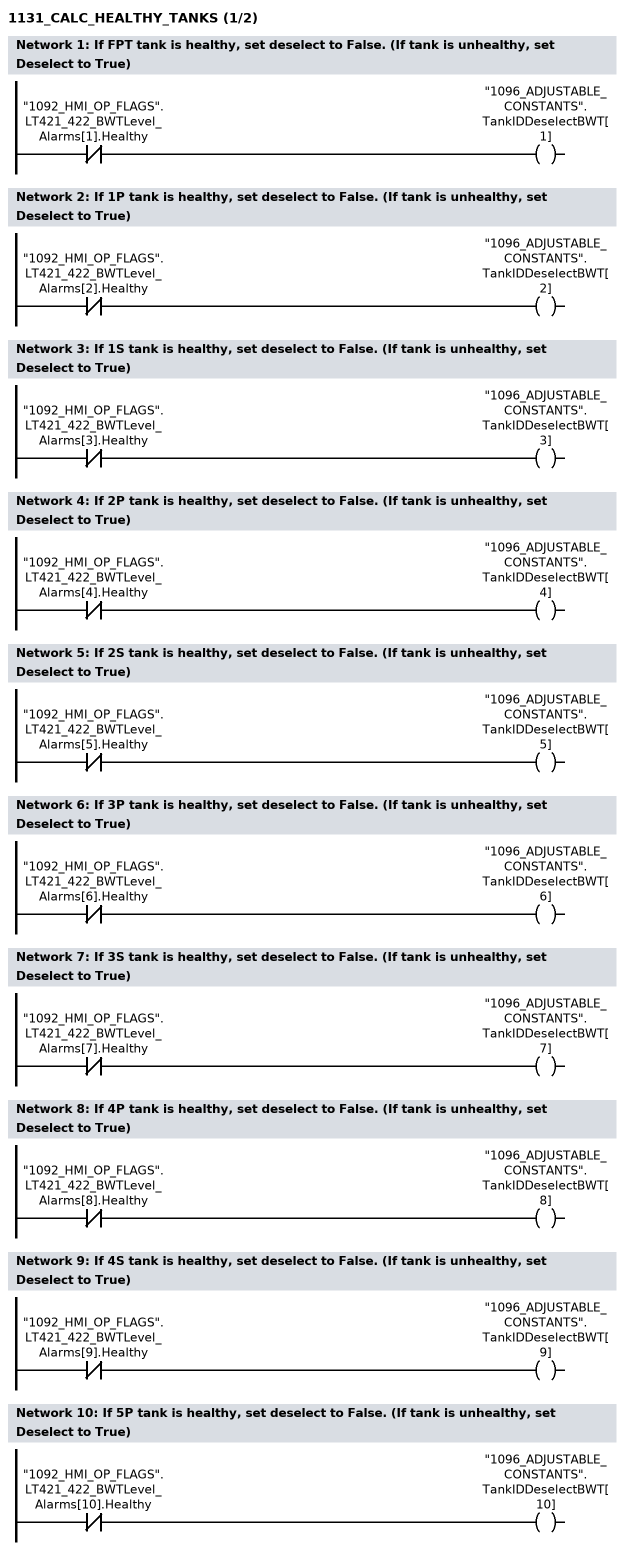
   RUNG wire#powerrail
      I_Contact( "1092_HMI_OP_FLAGS".LT421_422_BWTLevel_Alarms[1].Healthy )
      Coil( "1096_ADJUSTABLE_CONSTANTS".TankIDDeselectBWT[1] )
   END_RUNG
   // the same network as SCL:
   "1096_ADJUSTABLE_CONSTANTS".TankIDDeselectBWT[1] := NOT "1092_HMI_OP_FLAGS".LT421_422_BWTLevel_Alarms[1].Healthy;
END_REGION

REGION Network 2: If 1P tank is healthy, set deselect to False. (If tank is unhealthy, set Deselect to True)
   RUNG wire#powerrail
      I_Contact( "1092_HMI_OP_FLAGS".LT421_422_BWTLevel_Alarms[2].Healthy )
      Coil( "1096_ADJUSTABLE_CONSTANTS".TankIDDeselectBWT[2] )
   END_RUNG
   // the same network as SCL:
   "1096_ADJUSTABLE_CONSTANTS".TankIDDeselectBWT[2] := NOT "1092_HMI_OP_FLAGS".LT421_422_BWTLevel_Alarms[2].Healthy;
END_REGION

REGION Network 3: If 1S tank is healthy, set deselect to False. (If tank is unhealthy, set Deselect to True)
   RUNG wire#powerrail
      I_Contact( "1092_HMI_OP_FLAGS".LT421_422_BWTLevel_Alarms[3].Healthy )
      Coil( "1096_ADJUSTABLE_CONSTANTS".TankIDDeselectBWT[3] )
   END_RUNG
   // the same network as SCL:
   "1096_ADJUSTABLE_CONSTANTS".TankIDDeselectBWT[3] := NOT "1092_HMI_OP_FLAGS".LT421_422_BWTLevel_Alarms[3].Healthy;
END_REGION

REGION Network 4: If 2P tank is healthy, set deselect to False. (If tank is unhealthy, set Deselect to True)
   RUNG wire#powerrail
      I_Contact( "1092_HMI_OP_FLAGS".LT421_422_BWTLevel_Alarms[4].Healthy )
      Coil( "1096_ADJUSTABLE_CONSTANTS".TankIDDeselectBWT[4] )
   END_RUNG
   // the same network as SCL:
   "1096_ADJUSTABLE_CONSTANTS".TankIDDeselectBWT[4] := NOT "1092_HMI_OP_FLAGS".LT421_422_BWTLevel_Alarms[4].Healthy;
END_REGION

REGION Network 5: If 2S tank is healthy, set deselect to False. (If tank is unhealthy, set Deselect to True)
   RUNG wire#powerrail
      I_Contact( "1092_HMI_OP_FLAGS".LT421_422_BWTLevel_Alarms[5].Healthy )
      Coil( "1096_ADJUSTABLE_CONSTANTS".TankIDDeselectBWT[5] )
   END_RUNG
   // the same network as SCL:
   "1096_ADJUSTABLE_CONSTANTS".TankIDDeselectBWT[5] := NOT "1092_HMI_OP_FLAGS".LT421_422_BWTLevel_Alarms[5].Healthy;
END_REGION

REGION Network 6: If 3P tank is healthy, set deselect to False. (If tank is unhealthy, set Deselect to True)
   RUNG wire#powerrail
      I_Contact( "1092_HMI_OP_FLAGS".LT421_422_BWTLevel_Alarms[6].Healthy )
      Coil( "1096_ADJUSTABLE_CONSTANTS".TankIDDeselectBWT[6] )
   END_RUNG
   // the same network as SCL:
   "1096_ADJUSTABLE_CONSTANTS".TankIDDeselectBWT[6] := NOT "1092_HMI_OP_FLAGS".LT421_422_BWTLevel_Alarms[6].Healthy;
END_REGION

REGION Network 7: If 3S tank is healthy, set deselect to False. (If tank is unhealthy, set Deselect to True)
   RUNG wire#powerrail
      I_Contact( "1092_HMI_OP_FLAGS".LT421_422_BWTLevel_Alarms[7].Healthy )
      Coil( "1096_ADJUSTABLE_CONSTANTS".TankIDDeselectBWT[7] )
   END_RUNG
   // the same network as SCL:
   "1096_ADJUSTABLE_CONSTANTS".TankIDDeselectBWT[7] := NOT "1092_HMI_OP_FLAGS".LT421_422_BWTLevel_Alarms[7].Healthy;
END_REGION

REGION Network 8: If 4P tank is healthy, set deselect to False. (If tank is unhealthy, set Deselect to True)
   RUNG wire#powerrail
      I_Contact( "1092_HMI_OP_FLAGS".LT421_422_BWTLevel_Alarms[8].Healthy )
      Coil( "1096_ADJUSTABLE_CONSTANTS".TankIDDeselectBWT[8] )
   END_RUNG
   // the same network as SCL:
   "1096_ADJUSTABLE_CONSTANTS".TankIDDeselectBWT[8] := NOT "1092_HMI_OP_FLAGS".LT421_422_BWTLevel_Alarms[8].Healthy;
END_REGION

REGION Network 9: If 4S tank is healthy, set deselect to False. (If tank is unhealthy, set Deselect to True)
   RUNG wire#powerrail
      I_Contact( "1092_HMI_OP_FLAGS".LT421_422_BWTLevel_Alarms[9].Healthy )
      Coil( "1096_ADJUSTABLE_CONSTANTS".TankIDDeselectBWT[9] )
   END_RUNG
   // the same network as SCL:
   "1096_ADJUSTABLE_CONSTANTS".TankIDDeselectBWT[9] := NOT "1092_HMI_OP_FLAGS".LT421_422_BWTLevel_Alarms[9].Healthy;
END_REGION

REGION Network 10: If 5P tank is healthy, set deselect to False. (If tank is unhealthy, set Deselect to True)
   RUNG wire#powerrail
      I_Contact( "1092_HMI_OP_FLAGS".LT421_422_BWTLevel_Alarms[10].Healthy )
      Coil( "1096_ADJUSTABLE_CONSTANTS".TankIDDeselectBWT[10] )
   END_RUNG
   // the same network as SCL:
   "1096_ADJUSTABLE_CONSTANTS".TankIDDeselectBWT[10] := NOT "1092_HMI_OP_FLAGS".LT421_422_BWTLevel_Alarms[10].Healthy;
END_REGION

REGION Network 11: If 5S tank is healthy, set deselect to False. (If tank is unhealthy, set Deselect to True)
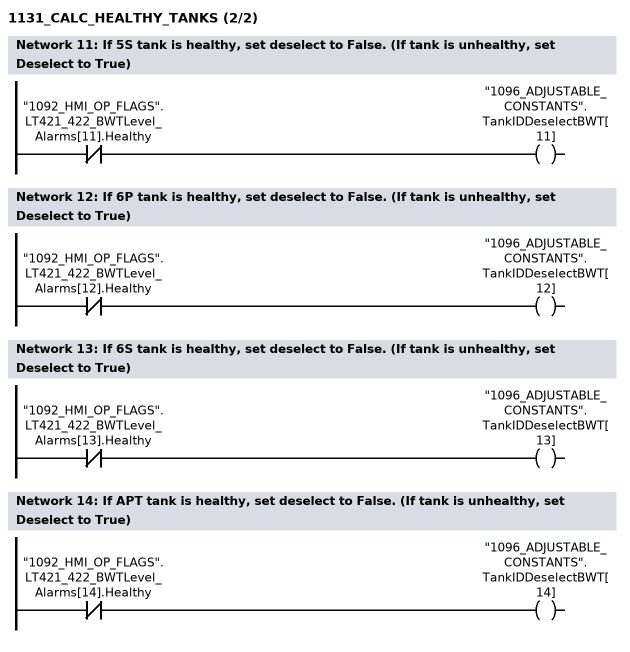
   RUNG wire#powerrail
      I_Contact( "1092_HMI_OP_FLAGS".LT421_422_BWTLevel_Alarms[11].Healthy )
      Coil( "1096_ADJUSTABLE_CONSTANTS".TankIDDeselectBWT[11] )
   END_RUNG
   // the same network as SCL:
   "1096_ADJUSTABLE_CONSTANTS".TankIDDeselectBWT[11] := NOT "1092_HMI_OP_FLAGS".LT421_422_BWTLevel_Alarms[11].Healthy;
END_REGION

REGION Network 12: If 6P tank is healthy, set deselect to False. (If tank is unhealthy, set Deselect to True)
   RUNG wire#powerrail
      I_Contact( "1092_HMI_OP_FLAGS".LT421_422_BWTLevel_Alarms[12].Healthy )
      Coil( "1096_ADJUSTABLE_CONSTANTS".TankIDDeselectBWT[12] )
   END_RUNG
   // the same network as SCL:
   "1096_ADJUSTABLE_CONSTANTS".TankIDDeselectBWT[12] := NOT "1092_HMI_OP_FLAGS".LT421_422_BWTLevel_Alarms[12].Healthy;
END_REGION

REGION Network 13: If 6S tank is healthy, set deselect to False. (If tank is unhealthy, set Deselect to True)
   RUNG wire#powerrail
      I_Contact( "1092_HMI_OP_FLAGS".LT421_422_BWTLevel_Alarms[13].Healthy )
      Coil( "1096_ADJUSTABLE_CONSTANTS".TankIDDeselectBWT[13] )
   END_RUNG
   // the same network as SCL:
   "1096_ADJUSTABLE_CONSTANTS".TankIDDeselectBWT[13] := NOT "1092_HMI_OP_FLAGS".LT421_422_BWTLevel_Alarms[13].Healthy;
END_REGION

REGION Network 14: If APT tank is healthy, set deselect to False. (If tank is unhealthy, set Deselect to True)
   RUNG wire#powerrail
      I_Contact( "1092_HMI_OP_FLAGS".LT421_422_BWTLevel_Alarms[14].Healthy )
      Coil( "1096_ADJUSTABLE_CONSTANTS".TankIDDeselectBWT[14] )
   END_RUNG
   // the same network as SCL:
   "1096_ADJUSTABLE_CONSTANTS".TankIDDeselectBWT[14] := NOT "1092_HMI_OP_FLAGS".LT421_422_BWTLevel_Alarms[14].Healthy;
END_REGION
END_FUNCTION

FUNCTION "1132_CALC_ACTIVE_TANKS" : Void   // FC1132, SCL
{ S7_Optimized_Access := 'TRUE' }
VERSION : 0.1
   VAR_TEMP
      Index : Int;
      NumberActiveTanks : Int;
   END_VAR
   VAR CONSTANT
      NumberOfTanks : Int := 14;
   END_VAR
BEGIN
   (*
       Calculate the number OF active tanks. With this data determine the HMI O/P flags:
       1. NoTanksActive (if no tanks are actively selected or healthy)
       2. The treatment time (the total treatment time of the vessel)
       3. Start IGG Warning Time (time flag to base IGG warnings on)
       4. VoyageLessThanTreatmentTime (error flag is the voyage will not be long enough to treat the tanks).
   *)

   #NumberActiveTanks := 0;

   FOR #Index := 1 TO #NumberOfTanks DO
       // For each tank that is not deselectable, force it to be active.
       IF NOT ("1096_ADJUSTABLE_CONSTANTS".TankIDDeselectBWT[#Index]) THEN
           "1096_ADJUSTABLE_CONSTANTS".TankIDActive[#Index] := TRUE;

       END_IF;
       // Check number of active tanks (either set in HMI, or by force above).
       IF "1096_ADJUSTABLE_CONSTANTS".TankIDActive[#Index] THEN
           #NumberActiveTanks += 1;
       END_IF;
   END_FOR;
   "1191_SYSTEM_VARIABLES".NumberOfActiveTanks := #NumberActiveTanks;

   // Push the no tanks active flag if calculated above.
   IF #NumberActiveTanks = 0 THEN
       "1092_HMI_OP_FLAGS".NoTanksActive := TRUE;
   ELSE
       "1092_HMI_OP_FLAGS".NoTanksActive := FALSE;
   END_IF;
END_FUNCTION

FUNCTION "1133_GTT_DETERMINE_EXCLUSIVITY" : Void   // FC1133, SCL
{ S7_Optimized_Access := 'TRUE' }
VERSION : 0.1
   VAR_INPUT
      TankID_InOperation : Int;
      DemandComplete : Bool;
   END_VAR
   VAR_IN_OUT
      GTT_Exclusivity : "GTT_EXCLUSIVITY";
   END_VAR
BEGIN
   (*
       Verify if the demand has been completed. If the demand is not yet complete,
       then keep this tank 'exclusive', i.e. do not allow another tank ID to begin 
       operating its GTT valve until this demand complete signal becomes True.
   *)

   IF NOT #DemandComplete THEN
       #GTT_Exclusivity.Tank_Exclusivity := TRUE;
       #GTT_Exclusivity.TankID_InOperation := #TankID_InOperation;
   ELSE
       #GTT_Exclusivity.Tank_Exclusivity := FALSE;
       #GTT_Exclusivity.TankID_InOperation := 0;
   END_IF;
END_FUNCTION

FUNCTION "1134_MOVE_TANKS_INGROUP_NEW_STATE" : Void   // FC1134, SCL
{ S7_Optimized_Access := 'TRUE' }
VERSION : 0.1
   VAR_INPUT
      State : "SYSTEM_STATES";
      NewState : Int;
   END_VAR
   VAR_IN_OUT
      TankData : Array[1..#NumberOfTanks] of "TANK_DATA";
   END_VAR
   VAR_TEMP
      Index : Int;
   END_VAR
   VAR CONSTANT
      NumberOfTanks : Int := 14;
   END_VAR
BEGIN
   (*
       For each tank, if it's in the current treatment group, 
       move it into the provided "NewState" state.
   *)
   FOR #Index := 1 TO #NumberOfTanks DO
       IF #TankData[#Index].AllocatedTreatmentGroup = #State.TreatmentGroup AND #TankData[#Index].Active THEN
           #TankData[#Index].TankState := #NewState;
       END_IF;
   END_FOR;
END_FUNCTION

FUNCTION "1135_VALVE_OPEN_CLOSE_TIME_SEL" : Time   // FC1135, SCL
{ S7_Optimized_Access := 'TRUE' }
VERSION : 0.1
   VAR_INPUT
      ValveType : Int;   // Valve Type. {0:NC,1:NO}
      ValveDemand : Bool;
      OpenTime : Time;
      CloseTime : Time;
   END_VAR
   VAR_TEMP
      SelectedTime : Time;
   END_VAR
   VAR CONSTANT
      Valve_NormallyClosed : Int := 0;
      Valve_NormallyOpen : Int := 1;
      Demand_Normal : Int := 0;
      Demand_Enable : Int := 1;
   END_VAR
BEGIN
   // Return the correct time for valve openning or closing based on whether
   // the valve is of type "Normally Open" or "Normally Closed" along with the
   // demand on the valve.
   CASE #ValveType OF
       #Valve_NormallyClosed:
           CASE BOOL_TO_INT(#ValveDemand) OF
               #Demand_Normal:
                   #SelectedTime := #CloseTime;
               #Demand_Enable:
                   #SelectedTime := #OpenTime;
           END_CASE;
       #Valve_NormallyOpen:
           CASE BOOL_TO_INT(#ValveDemand) OF
               #Demand_Normal:
                   #SelectedTime := #OpenTime;
               #Demand_Enable:
                   #SelectedTime := #CloseTime;
           END_CASE;
   END_CASE;

   #"1135_VALVE_OPEN_CLOSE_TIME_SEL" := #SelectedTime;
END_FUNCTION

FUNCTION "1136_CALC_NEXT_TREATMENT_GROUP" : Int   // FC1136, SCL
{ S7_Optimized_Access := 'TRUE' }
VERSION : 0.1
   VAR_INPUT
      State : "SYSTEM_STATES";
      NumberOfTreatmentGroups : Int;
      TankData : Array[1..#NumberOfTanks] of "TANK_DATA";
   END_VAR
   VAR_TEMP
      NextTreatmentGroupCalc : Int;
      NextTreatmentGroupFound : Bool;
      TreatmentGroupContainsActiveTank : Bool;
      Index : Int;
   END_VAR
   VAR CONSTANT
      NumberOfTanks : Int := 14;
   END_VAR
BEGIN
   // Return the next treatment group ID which contains active tanks.
   // Return a -1 if there are no further active tanks, or this is the greatest tank ID.
   #NextTreatmentGroupFound := False;
   #NextTreatmentGroupCalc := #State.TreatmentGroup + 1;

   IF #NextTreatmentGroupCalc <= #NumberOfTreatmentGroups THEN
       WHILE NOT #NextTreatmentGroupFound DO
           // Another treatment group to go, check if there are active tanks in the next group.
           #TreatmentGroupContainsActiveTank := False;
           FOR #Index := 1 TO #NumberOfTanks DO
               IF #TankData[#Index].AllocatedTreatmentGroup = #NextTreatmentGroupCalc AND "1096_ADJUSTABLE_CONSTANTS".TankIDActive[#Index] = True THEN
                   #TreatmentGroupContainsActiveTank := True;
               END_IF;
           END_FOR;
           IF #TreatmentGroupContainsActiveTank = True THEN
               // A treatment group has been found.
               #NextTreatmentGroupFound := True;
           ELSE
               // A treatment group was not found on this cycle, check if there are more treatment groups to go.
               IF #NextTreatmentGroupCalc + 1 <= #NumberOfTreatmentGroups THEN
                   #NextTreatmentGroupCalc += 1;
               ELSE
                   // No treatment groups remain, return -1.
                   #NextTreatmentGroupCalc := -1;
                   #NextTreatmentGroupFound := True;
               END_IF;
           END_IF;
       END_WHILE;
   ELSE
       // This is the last treatment group, return a -1 to show that there are no further groups.
       #NextTreatmentGroupCalc := -1;
   END_IF;

   #"1136_CALC_NEXT_TREATMENT_GROUP" := #NextTreatmentGroupCalc;
END_FUNCTION

// folder: 1000 - 1999 BWT System Control/1130 - 1159 Support Functions/1150 - 1159 Next Stage Checks

FUNCTION "1150_NEXT_STAGE_CHECK_GTT" : "ALARM_DEMAND_RTN"   // FC1150, SCL
{ S7_Optimized_Access := 'TRUE' }
VERSION : 0.1
   VAR_INPUT
      AlarmState : Int;   // State system should move to in the event of an alarm being raised (Normally State_Shutdown)
      GTT_OUT : "VALVE_GTT_OUT";
      TankData : Array[1..#NumberOfTanks] of "TANK_DATA";
   END_VAR
   VAR_IN_OUT
      State : "SYSTEM_STATES";
   END_VAR
   VAR_TEMP
      Index : Int;
      NextStageCheck : "ALARM_DEMAND_RTN";
   END_VAR
   VAR CONSTANT
      NumberOfTanks : Int := 14;
   END_VAR
BEGIN
   (*
       Function to check whether the treatment group is ready to move to the next stage
       This specifically checks the GTT completion and will return the demand complete
       only once all active tanks have completed GTT actuation actions.
   *)

   #NextStageCheck.Demand_Complete := True;
   #NextStageCheck.Alarm_Active := False;

   FOR #Index := 1 TO #NumberOfTanks DO
       IF #TankData[#Index].AllocatedTreatmentGroup = #State.TreatmentGroup AND #TankData[#Index].Active THEN
           IF NOT (#GTT_OUT.GTT_DemandsCompleted[#Index]) THEN
               #NextStageCheck.Demand_Complete := False;
           END_IF;
           IF #GTT_OUT.GTT_Alarms[#Index] THEN
               #NextStageCheck.Alarm_Active := True;
           END_IF;
       END_IF;
   END_FOR;

   IF #NextStageCheck.Alarm_Active THEN
       #State.System := #AlarmState;
   END_IF;

   #"1150_NEXT_STAGE_CHECK_GTT" := #NextStageCheck;
END_FUNCTION

FUNCTION "1151_NEXT_STAGE_CHECK_PVV" : "ALARM_DEMAND_RTN"   // FC1151, SCL
{ S7_Optimized_Access := 'TRUE' }
VERSION : 0.1
   VAR_INPUT
      AlarmState : Int;   // State system should move to in the event of an alarm being raised (Normally State_Shutdown)
      PVVX_OUT : "VALVE_PVVX_OUT";
      TankData : Array[1..#NumberOfTanks] of "TANK_DATA";
   END_VAR
   VAR_IN_OUT
      State : "SYSTEM_STATES";
   END_VAR
   VAR_TEMP
      Index : Int;
      NextStageCheck : "ALARM_DEMAND_RTN";
   END_VAR
   VAR CONSTANT
      NumberOfTanks : Int := 14;
   END_VAR
BEGIN
   (*
       Function to check whether the treatment group is ready to move to the next stage
       This specifically checks the Vent A/B completion and will return the demand complete
       only once all active tanks have completed Vent A/B actuation actions.
   *)

   #NextStageCheck.Demand_Complete := True;
   #NextStageCheck.Alarm_Active := False;

   FOR #Index := 1 TO #NumberOfTanks DO
       IF #TankData[#Index].AllocatedTreatmentGroup = #State.TreatmentGroup AND #TankData[#Index].Active THEN
           IF NOT (#PVVX_OUT.PVVA_DemandsCompleted[#Index] OR #PVVX_OUT.PVVB_DemandsCompleted[#Index]) THEN
               #NextStageCheck.Demand_Complete := False;
           END_IF;
           IF (#PVVX_OUT.PVVA_Alarms[#Index] OR #PVVX_OUT.PVVB_Alarms[#Index]) THEN
               #NextStageCheck.Alarm_Active := True;
           END_IF;
       END_IF;
   END_FOR;

   IF #NextStageCheck.Alarm_Active THEN
       #State.System := #AlarmState;
   END_IF;

   #"1151_NEXT_STAGE_CHECK_PVV" := #NextStageCheck;
END_FUNCTION

FUNCTION "1152_NEXT_STAGE_CHECK_TIMER" : "ALARM_DEMAND_RTN"   // FC1152, SCL
{ S7_Optimized_Access := 'TRUE' }
VERSION : 0.1
   VAR_INPUT
      AlarmState : Int;   // State system should move to in the event of an alarm being raised (Normally State_Shutdown)
      TankData : Array[1..#NumberOfTanks] of "TANK_DATA";
   END_VAR
   VAR_IN_OUT
      State : "SYSTEM_STATES";
   END_VAR
   VAR_TEMP
      Index : Int;
      NextStageCheck : "ALARM_DEMAND_RTN";
   END_VAR
   VAR CONSTANT
      NumberOfTanks : Int := 14;
   END_VAR
BEGIN
   (*
       Function to check whether the treatment group is ready to move to the next stage
       This specifically checks the the timer of a tank (xx-Dwell) completion and will return
       the demand complete only once all active tanks have completed their timeouts, depending
       on the overall system state, this is a multi-function block call
   *)

   #NextStageCheck.Demand_Complete := True;
   #NextStageCheck.Alarm_Active := False;

   FOR #Index := 1 TO #NumberOfTanks DO
       IF #TankData[#Index].AllocatedTreatmentGroup = #State.TreatmentGroup AND #TankData[#Index].Active THEN
           IF NOT (#TankData[#Index].Timer_Complete) THEN
               #NextStageCheck.Demand_Complete := False;
           END_IF;
       END_IF;
   END_FOR;

   IF #NextStageCheck.Alarm_Active THEN
       #State.System := #AlarmState;
   END_IF;

   #"1152_NEXT_STAGE_CHECK_TIMER" := #NextStageCheck;
END_FUNCTION

FUNCTION "1153_NEXT_STAGE_CHECK_XEOX" : "ALARM_DEMAND_RTN"   // FC1153, SCL
{ S7_Optimized_Access := 'TRUE' }
VERSION : 0.1
   VAR_INPUT
      AlarmState : Int;   // State system should move to in the event of an alarm being raised (Normally State_Shutdown)
      TankData : Array[1..#NumberOfTanks] of "TANK_DATA";
   END_VAR
   VAR_IN_OUT
      State : "SYSTEM_STATES";
   END_VAR
   VAR_TEMP
      Index : Int;
      NextStageCheck : "ALARM_DEMAND_RTN";
   END_VAR
   VAR CONSTANT
      NumberOfTanks : Int := 14;
   END_VAR
BEGIN
   (*
       Function to check whether the treatment group is ready to move to the next stage
       This specifically checks the the ReOx/DeOx of a tank completion and will return
       the demand complete only once all active tanks have completed ReOx or DeOx, depending
       on the overall system state, this is a multi-function block call
   *)

   #NextStageCheck.Demand_Complete := True;
   #NextStageCheck.Alarm_Active := False;

   FOR #Index := 1 TO #NumberOfTanks DO
       IF #TankData[#Index].AllocatedTreatmentGroup = #State.TreatmentGroup AND #TankData[#Index].Active THEN
           IF NOT (#TankData[#Index].XeOx_Complete) THEN
               #NextStageCheck.Demand_Complete := False;
           END_IF;
       END_IF;
   END_FOR;

   IF #NextStageCheck.Alarm_Active THEN
       #State.System := #AlarmState;
   END_IF;

   #"1153_NEXT_STAGE_CHECK_XEOX" := #NextStageCheck;
END_FUNCTION

// folder: 1000 - 1999 BWT System Control/1600 - 1999 Standard FB's

FUNCTION_BLOCK "1604_DEMAND_AND_CHECK"   // FB1604, LAD
TITLE = Valve Check
{ S7_Optimized_Access := 'TRUE' }
AUTHOR : JRS
VERSION : 0.1
// Demand and check an NO or NC valve.
   VAR_INPUT
      DemandIn : Bool;   // Demand
      NO_Type : Bool;   // Valve type = open without demand
      NC_Type : Bool;   // Valve type = closed without demand
      ValveMoveTime : LTime := LT#1s;   // Maximum movement time
      ValveOpenStatus : Bool;   // Valve open confirmed
      ValveClsdStatus : Bool;   // Valve closed confirmed
   END_VAR
   VAR_OUTPUT
      DemandOut : Bool;   // Demand feedthrough from DemandIn
      DemandComplete : Bool;   // Valve has completed movement
      Alarm : Bool;   // Valve is faulty
   END_VAR
   VAR RETAIN
      Reset : Bool := True;
      Healthy : Bool;   // Valve is healthy
      Config_Error : Bool;   // Configuration error
      Sensor_Fault : Bool;   // Sensor conflicts
      TRAVEL_TIME : TONR_LTIME;
   END_VAR
BEGIN

REGION Network 1: Configuration Error
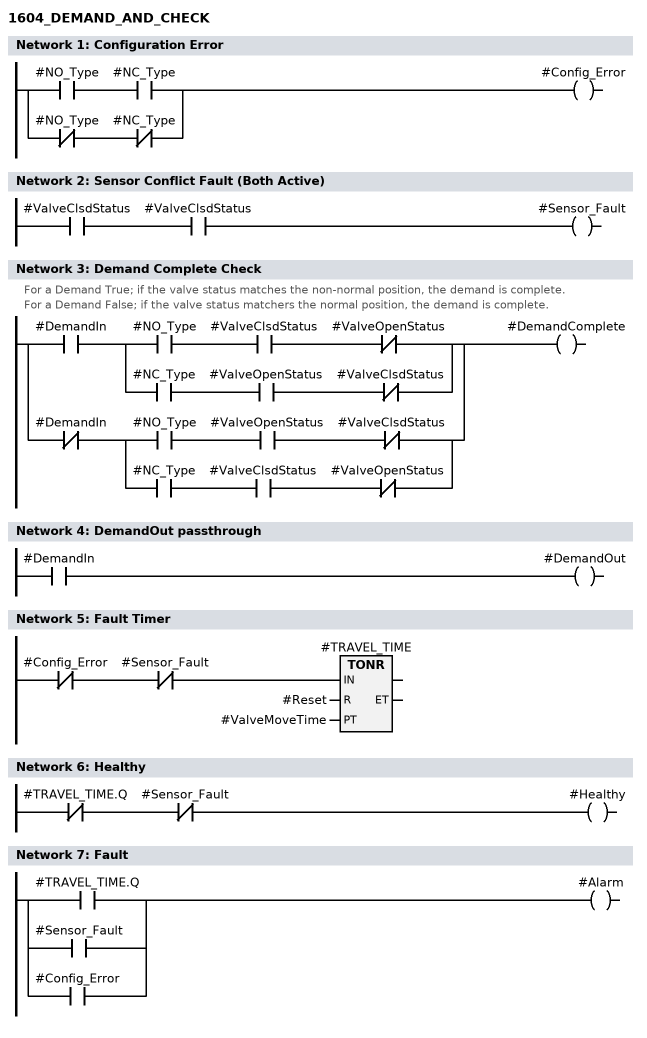
   RUNG wire#powerrail
      Contact( #NO_Type )
      Contact( #NC_Type )
      wire#w1
      Coil( #Config_Error )
   END_RUNG
   RUNG wire#powerrail
      I_Contact( #NO_Type )
      I_Contact( #NC_Type )
   END_RUNG wire#w1
   // the same network as SCL:
   #Config_Error := (#NO_Type AND #NC_Type) OR (NOT #NO_Type AND NOT #NC_Type);
END_REGION

REGION Network 2: Sensor Conflict Fault (Both Active)
   RUNG wire#powerrail
      Contact( #ValveClsdStatus )
      Contact( #ValveClsdStatus )
      Coil( #Sensor_Fault )
   END_RUNG
   // the same network as SCL:
   #Sensor_Fault := #ValveClsdStatus AND #ValveClsdStatus;
END_REGION

REGION Network 3: Demand Complete Check
   // For a Demand True; if the valve status matches the non-normal position, the demand is complete.
   // For a Demand False; if the valve status matchers the normal position, the demand is complete.
   RUNG wire#powerrail
      Contact( #DemandIn )
      wire#w1
      Contact( #NO_Type )
      Contact( #ValveClsdStatus )
      I_Contact( #ValveOpenStatus )
      wire#w2
      Coil( #DemandComplete )
   END_RUNG
   RUNG wire#w1
      Contact( #NC_Type )
      Contact( #ValveOpenStatus )
      I_Contact( #ValveClsdStatus )
   END_RUNG wire#w2
   RUNG wire#powerrail
      I_Contact( #DemandIn )
      wire#w3
      Contact( #NO_Type )
      Contact( #ValveOpenStatus )
      I_Contact( #ValveClsdStatus )
   END_RUNG wire#w2
   RUNG wire#w3
      Contact( #NC_Type )
      Contact( #ValveClsdStatus )
      I_Contact( #ValveOpenStatus )
   END_RUNG wire#w2
   // the same network as SCL:
   #DemandComplete := (#DemandIn AND ((#NO_Type AND #ValveClsdStatus AND NOT #ValveOpenStatus) OR (#NC_Type AND #ValveOpenStatus AND NOT #ValveClsdStatus))) OR (NOT #DemandIn AND ((#NO_Type AND #ValveOpenStatus AND NOT #ValveClsdStatus) OR (#NC_Type AND #ValveClsdStatus AND NOT #ValveOpenStatus)));
END_REGION

REGION Network 4: DemandOut passthrough
   RUNG wire#powerrail
      Contact( #DemandIn )
      Coil( #DemandOut )
   END_RUNG
   // the same network as SCL:
   #DemandOut := #DemandIn;
END_REGION

REGION Network 5: Fault Timer
   #TRAVEL_TIME(IN := NOT #Config_Error AND NOT #Sensor_Fault, R := #Reset, PT := #ValveMoveTime);   // TONR
END_REGION

REGION Network 6: Healthy
   RUNG wire#powerrail
      I_Contact( #TRAVEL_TIME.Q )
      I_Contact( #Sensor_Fault )
      Coil( #Healthy )
   END_RUNG
   // the same network as SCL:
   #Healthy := NOT #TRAVEL_TIME.Q AND NOT #Sensor_Fault;
END_REGION

REGION Network 7: Fault
   RUNG wire#powerrail
      Contact( #TRAVEL_TIME.Q )
      wire#w1
      Coil( #Alarm )
   END_RUNG
   RUNG wire#powerrail
      Contact( #Sensor_Fault )
   END_RUNG wire#w1
   RUNG wire#powerrail
      Contact( #Config_Error )
   END_RUNG wire#w1
   // the same network as SCL:
   #Alarm := #TRAVEL_TIME.Q OR #Sensor_Fault OR #Config_Error;
END_REGION
END_FUNCTION_BLOCK

FUNCTION "1601_ANALOGUE_HEALTH_ALLTRIPS" : Void   // FC1601, LAD
{ S7_Optimized_Access := 'TRUE' }
VERSION : 0.1
   VAR_INPUT
      InputSignal : Real;   // Analogue sensor value
      InputMinimum : Real;   // Minimum sensor value
      InputMaximum : Real;   // Maximum sensor value
      InputSetpointLowLow : Real;   // Low low setpoint value for sensor
      InputSetpointLow : Real;   // Low setpoint value for sensor
      InputSetpointHigh : Real;   // High setpoint value for sensor
      InputSetpointHighHigh : Real;   // High high setpoint value for sensor
   END_VAR
   VAR_OUTPUT
      SensorHealthOut : Bool;   // Boolean health status
      LowLowAlarmOut : Bool;   // Boolean for low low alarm
      LowWarningOut : Bool;   // Boolean for low warning
      HighWarningOut : Bool;   // Boolean for high warning
      HighHighAlarmOut : Bool;   // Boolean for high high alarm
   END_VAR
BEGIN

REGION Network 1: Boolean health status
   // Determine SensorHealthOut (health status) dependent on input signal from sensor compared to setpoints. [GEN-05]
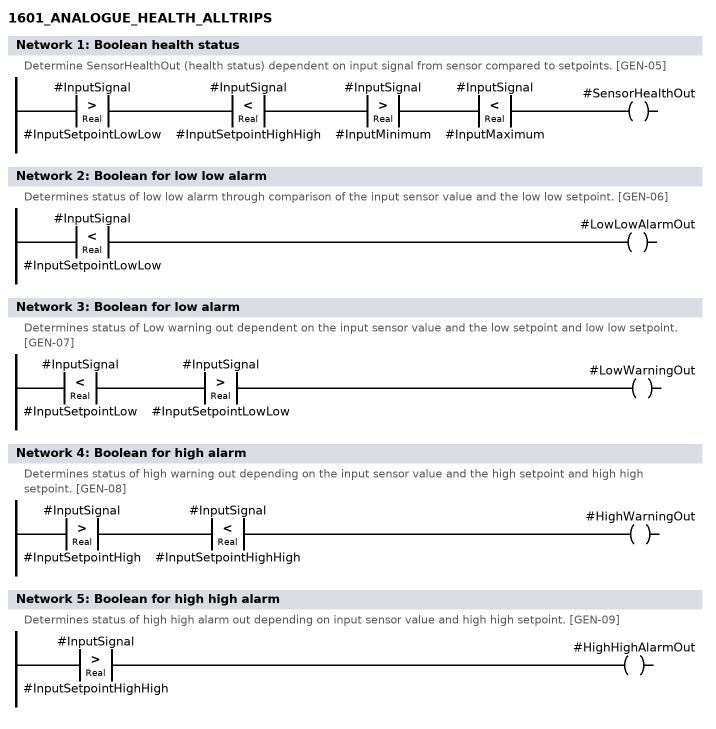
   RUNG wire#powerrail
      { S7_Templates := "SrcType := Real" } GT_Contact(in1 := #InputSignal, in2 := #InputSetpointLowLow)
      { S7_Templates := "SrcType := Real" } LT_Contact(in1 := #InputSignal, in2 := #InputSetpointHighHigh)
      { S7_Templates := "SrcType := Real" } GT_Contact(in1 := #InputSignal, in2 := #InputMinimum)
      { S7_Templates := "SrcType := Real" } LT_Contact(in1 := #InputSignal, in2 := #InputMaximum)
      Coil( #SensorHealthOut )
   END_RUNG
   // the same network as SCL:
   #SensorHealthOut := (#InputSignal > #InputSetpointLowLow) AND (#InputSignal < #InputSetpointHighHigh) AND (#InputSignal > #InputMinimum) AND (#InputSignal < #InputMaximum);
END_REGION

REGION Network 2: Boolean for low low alarm
   // Determines status of low low alarm through comparison of the input sensor value and the low low setpoint. [GEN-06]
   RUNG wire#powerrail
      { S7_Templates := "SrcType := Real" } LT_Contact(in1 := #InputSignal, in2 := #InputSetpointLowLow)
      Coil( #LowLowAlarmOut )
   END_RUNG
   // the same network as SCL:
   #LowLowAlarmOut := #InputSignal < #InputSetpointLowLow;
END_REGION

REGION Network 3: Boolean for low alarm
   // Determines status of Low warning out dependent on the input sensor value and the low setpoint and low low setpoint. [GEN-07]
   RUNG wire#powerrail
      { S7_Templates := "SrcType := Real" } LT_Contact(in1 := #InputSignal, in2 := #InputSetpointLow)
      { S7_Templates := "SrcType := Real" } GT_Contact(in1 := #InputSignal, in2 := #InputSetpointLowLow)
      Coil( #LowWarningOut )
   END_RUNG
   // the same network as SCL:
   #LowWarningOut := (#InputSignal < #InputSetpointLow) AND (#InputSignal > #InputSetpointLowLow);
END_REGION

REGION Network 4: Boolean for high alarm
   // Determines status of high warning out depending on the input sensor value and the high setpoint and high high setpoint. [GEN-08]
   RUNG wire#powerrail
      { S7_Templates := "SrcType := Real" } GT_Contact(in1 := #InputSignal, in2 := #InputSetpointHigh)
      { S7_Templates := "SrcType := Real" } LT_Contact(in1 := #InputSignal, in2 := #InputSetpointHighHigh)
      Coil( #HighWarningOut )
   END_RUNG
   // the same network as SCL:
   #HighWarningOut := (#InputSignal > #InputSetpointHigh) AND (#InputSignal < #InputSetpointHighHigh);
END_REGION

REGION Network 5: Boolean for high high alarm
   // Determines status of high high alarm out depending on input sensor value and high high setpoint. [GEN-09]
   RUNG wire#powerrail
      { S7_Templates := "SrcType := Real" } GT_Contact(in1 := #InputSignal, in2 := #InputSetpointHighHigh)
      Coil( #HighHighAlarmOut )
   END_RUNG
   // the same network as SCL:
   #HighHighAlarmOut := #InputSignal > #InputSetpointHighHigh;
END_REGION
END_FUNCTION

FUNCTION "1602_DIGITAL_HEALTH" : Void   // FC1602, LAD
{ S7_Optimized_Access := 'TRUE' }
VERSION : 0.1
   VAR_INPUT
      InputSignal : Bool;   // Digital sensor value
      InputTripLevel : Bool;   // Nature of trip value
   END_VAR
   VAR_OUTPUT
      SensorHealthOut : Bool;   // Boolean health status
      AlarmOut : Bool;   // Boolean alarm status
   END_VAR
BEGIN

REGION Network 1: Boolean alarm status
   // Sensor is healthy only if its input is high for a low level trip or low for a high level trip. [GEN-17]
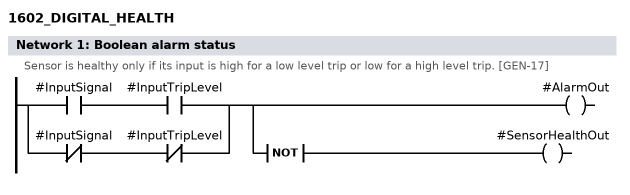
   RUNG wire#powerrail
      Contact( #InputSignal )
      Contact( #InputTripLevel )
      wire#w1
      Coil( #AlarmOut )
   END_RUNG
   RUNG wire#powerrail
      I_Contact( #InputSignal )
      I_Contact( #InputTripLevel )
   END_RUNG wire#w1
   RUNG wire#w1
      Not()
      Coil( #SensorHealthOut )
   END_RUNG
   // the same network as SCL:
   #AlarmOut := (#InputSignal AND #InputTripLevel) OR (NOT #InputSignal AND NOT #InputTripLevel);
   #SensorHealthOut := NOT #AlarmOut;
END_REGION
END_FUNCTION

FUNCTION "1603_VALVE_STATE" : Void   // FC1603, SCL
{ S7_Optimized_Access := 'TRUE' }
VERSION : 0.1
   VAR_INPUT
      InputLimitSwitchOpen : Bool;   // True indicates that the limit switch is closed.
      InputLimitSwitchClosed : Bool;   // True indicates that the limit switch is closed.
   END_VAR
   VAR_OUTPUT
      Open : Bool;   // Valve Open Status
      Closed : Bool;   // Valve Closed Status
      Moving : Bool;   // Valve Moving Status
      Fault : Bool;   // Valve Fault Status
   END_VAR
BEGIN
   (*
   This function dictates the Open/Closed/Moving/Fault status of the valve
   depending on the inputs Limit Switch Open, Limit Switch closed.
   [GEN-38]
   *)

   IF ((#InputLimitSwitchOpen = TRUE) AND (#InputLimitSwitchClosed = FALSE)) THEN
       #Open := TRUE;
       #Closed := FALSE;
       #Moving := FALSE;
       #Fault := FALSE;
   ELSIF ((#InputLimitSwitchOpen = TRUE) AND (#InputLimitSwitchClosed = TRUE)) THEN
       #Open := FALSE;
       #Closed := FALSE;
       #Moving := FALSE;
       #Fault := TRUE;
   ELSIF ((#InputLimitSwitchOpen = FALSE) AND (#InputLimitSwitchClosed = FALSE)) THEN
       #Open := FALSE;
       #Closed := FALSE;
       #Moving := TRUE;
       #Fault := FALSE;
   ELSE
       #Open := FALSE;
       #Closed := TRUE;
       #Moving := FALSE;
       #Fault := FALSE;
   END_IF;
END_FUNCTION

// folder: 20 - 49 RIO & Processing

FUNCTION "20_RIO_Input_Processing" : Void   // FC20, LAD
TITLE = RIO Input Processing
{ S7_Optimized_Access := 'TRUE' }
AUTHOR : JRS
VERSION : 0.1
// To call input processing blocks in logical order
BEGIN

REGION Network 1: RIO Digital Input Processing - Rack 1
   // To process raw inputs prior to code use
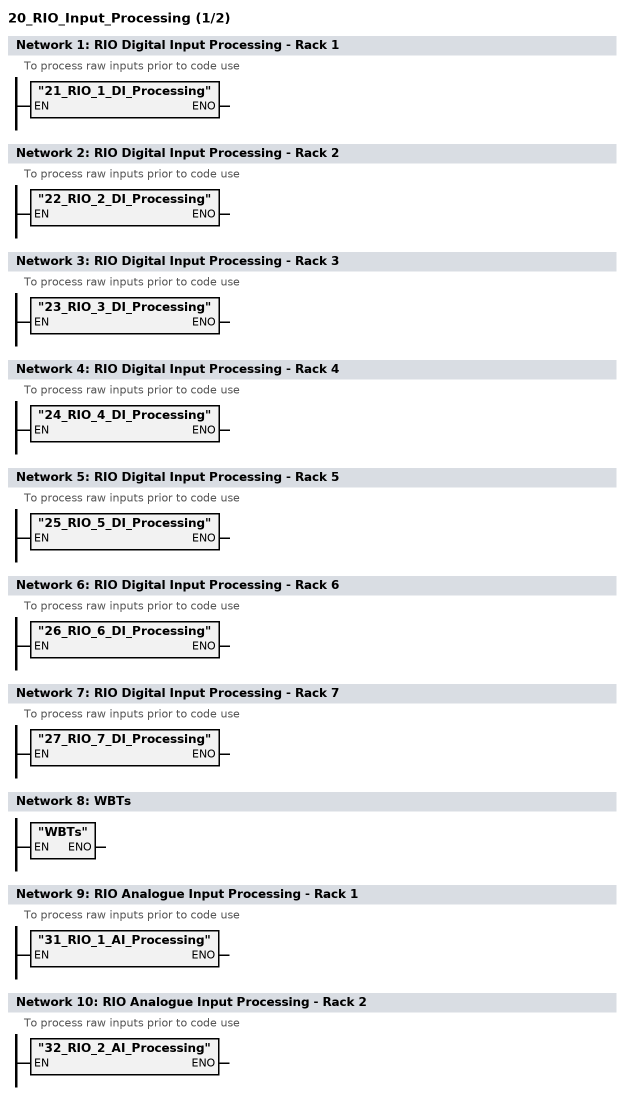
   RUNG wire#powerrail
      "21_RIO_1_DI_Processing"()
   END_RUNG
   // the same network as SCL:
   "21_RIO_1_DI_Processing"();
END_REGION

REGION Network 2: RIO Digital Input Processing - Rack 2
   // To process raw inputs prior to code use
   RUNG wire#powerrail
      "22_RIO_2_DI_Processing"()
   END_RUNG
   // the same network as SCL:
   "22_RIO_2_DI_Processing"();
END_REGION

REGION Network 3: RIO Digital Input Processing - Rack 3
   // To process raw inputs prior to code use
   RUNG wire#powerrail
      "23_RIO_3_DI_Processing"()
   END_RUNG
   // the same network as SCL:
   "23_RIO_3_DI_Processing"();
END_REGION

REGION Network 4: RIO Digital Input Processing - Rack 4
   // To process raw inputs prior to code use
   RUNG wire#powerrail
      "24_RIO_4_DI_Processing"()
   END_RUNG
   // the same network as SCL:
   "24_RIO_4_DI_Processing"();
END_REGION

REGION Network 5: RIO Digital Input Processing - Rack 5
   // To process raw inputs prior to code use
   RUNG wire#powerrail
      "25_RIO_5_DI_Processing"()
   END_RUNG
   // the same network as SCL:
   "25_RIO_5_DI_Processing"();
END_REGION

REGION Network 6: RIO Digital Input Processing - Rack 6
   // To process raw inputs prior to code use
   RUNG wire#powerrail
      "26_RIO_6_DI_Processing"()
   END_RUNG
   // the same network as SCL:
   "26_RIO_6_DI_Processing"();
END_REGION

REGION Network 7: RIO Digital Input Processing - Rack 7
   // To process raw inputs prior to code use
   RUNG wire#powerrail
      "27_RIO_7_DI_Processing"()
   END_RUNG
   // the same network as SCL:
   "27_RIO_7_DI_Processing"();
END_REGION

REGION Network 8: WBTs
   RUNG wire#powerrail
      "WBTs"()
   END_RUNG
   // the same network as SCL:
   "WBTs"();
END_REGION

REGION Network 9: RIO Analogue Input Processing - Rack 1
   // To process raw inputs prior to code use
   RUNG wire#powerrail
      "31_RIO_1_AI_Processing"()
   END_RUNG
   // the same network as SCL:
   "31_RIO_1_AI_Processing"();
END_REGION

REGION Network 10: RIO Analogue Input Processing - Rack 2
   // To process raw inputs prior to code use
   RUNG wire#powerrail
      "32_RIO_2_AI_Processing"()
   END_RUNG
   // the same network as SCL:
   "32_RIO_2_AI_Processing"();
END_REGION

REGION Network 11: RIO Analogue Input Processing - Rack 3
   // To process raw inputs prior to code use
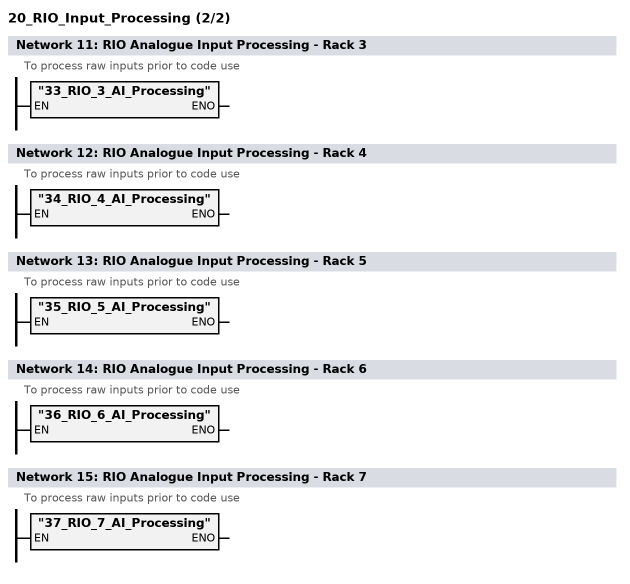
   RUNG wire#powerrail
      "33_RIO_3_AI_Processing"()
   END_RUNG
   // the same network as SCL:
   "33_RIO_3_AI_Processing"();
END_REGION

REGION Network 12: RIO Analogue Input Processing - Rack 4
   // To process raw inputs prior to code use
   RUNG wire#powerrail
      "34_RIO_4_AI_Processing"()
   END_RUNG
   // the same network as SCL:
   "34_RIO_4_AI_Processing"();
END_REGION

REGION Network 13: RIO Analogue Input Processing - Rack 5
   // To process raw inputs prior to code use
   RUNG wire#powerrail
      "35_RIO_5_AI_Processing"()
   END_RUNG
   // the same network as SCL:
   "35_RIO_5_AI_Processing"();
END_REGION

REGION Network 14: RIO Analogue Input Processing - Rack 6
   // To process raw inputs prior to code use
   RUNG wire#powerrail
      "36_RIO_6_AI_Processing"()
   END_RUNG
   // the same network as SCL:
   "36_RIO_6_AI_Processing"();
END_REGION

REGION Network 15: RIO Analogue Input Processing - Rack 7
   // To process raw inputs prior to code use
   RUNG wire#powerrail
      "37_RIO_7_AI_Processing"()
   END_RUNG
   // the same network as SCL:
   "37_RIO_7_AI_Processing"();
END_REGION
END_FUNCTION

FUNCTION "21_RIO_1_DI_Processing" : Void   // FC21, LAD
TITLE = RIO Rack Digital Input Processing (Tank 1 = FPT, Tank 2 = 1P, Tank 3 = 1S)
{ S7_Optimized_Access := 'TRUE' }
AUTHOR : JRS
VERSION : 0.1
// To process raw inputs prior to code use
BEGIN

REGION Network 1: I0.0 - Gas To Tank Valve Feedback Open (CV-422)
   // True = OPEN, False = NOT
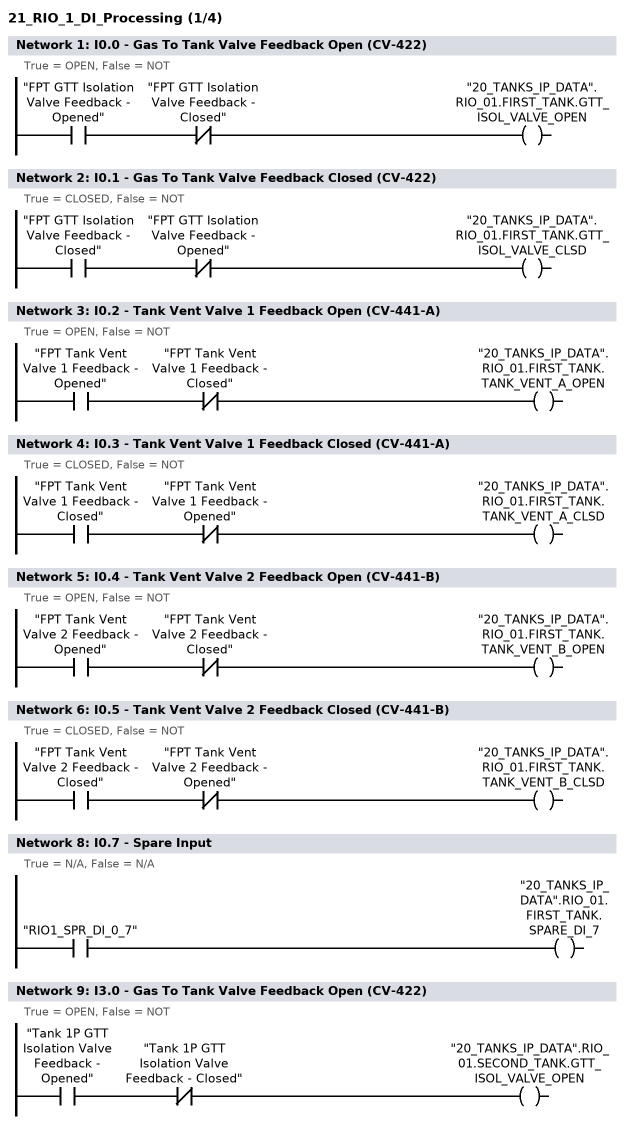
   RUNG wire#powerrail
      Contact( "FPT GTT Isolation Valve Feedback - Opened" )
      I_Contact( "FPT GTT Isolation Valve Feedback - Closed" )
      Coil( "20_TANKS_IP_DATA".RIO_01.FIRST_TANK.GTT_ISOL_VALVE_OPEN )
   END_RUNG
   // the same network as SCL:
   "20_TANKS_IP_DATA".RIO_01.FIRST_TANK.GTT_ISOL_VALVE_OPEN := "FPT GTT Isolation Valve Feedback - Opened" AND NOT "FPT GTT Isolation Valve Feedback - Closed";
END_REGION

REGION Network 2: I0.1 - Gas To Tank Valve Feedback Closed (CV-422)
   // True = CLOSED, False = NOT
   RUNG wire#powerrail
      Contact( "FPT GTT Isolation Valve Feedback - Closed" )
      I_Contact( "FPT GTT Isolation Valve Feedback - Opened" )
      Coil( "20_TANKS_IP_DATA".RIO_01.FIRST_TANK.GTT_ISOL_VALVE_CLSD )
   END_RUNG
   // the same network as SCL:
   "20_TANKS_IP_DATA".RIO_01.FIRST_TANK.GTT_ISOL_VALVE_CLSD := "FPT GTT Isolation Valve Feedback - Closed" AND NOT "FPT GTT Isolation Valve Feedback - Opened";
END_REGION

REGION Network 3: I0.2 - Tank Vent Valve 1 Feedback Open (CV-441-A)
   // True = OPEN, False = NOT
   RUNG wire#powerrail
      Contact( "FPT Tank Vent Valve 1 Feedback - Opened" )
      I_Contact( "FPT Tank Vent Valve 1 Feedback - Closed" )
      Coil( "20_TANKS_IP_DATA".RIO_01.FIRST_TANK.TANK_VENT_A_OPEN )
   END_RUNG
   // the same network as SCL:
   "20_TANKS_IP_DATA".RIO_01.FIRST_TANK.TANK_VENT_A_OPEN := "FPT Tank Vent Valve 1 Feedback - Opened" AND NOT "FPT Tank Vent Valve 1 Feedback - Closed";
END_REGION

REGION Network 4: I0.3 - Tank Vent Valve 1 Feedback Closed (CV-441-A)
   // True = CLOSED, False = NOT
   RUNG wire#powerrail
      Contact( "FPT Tank Vent Valve 1 Feedback - Closed" )
      I_Contact( "FPT Tank Vent Valve 1 Feedback - Opened" )
      Coil( "20_TANKS_IP_DATA".RIO_01.FIRST_TANK.TANK_VENT_A_CLSD )
   END_RUNG
   // the same network as SCL:
   "20_TANKS_IP_DATA".RIO_01.FIRST_TANK.TANK_VENT_A_CLSD := "FPT Tank Vent Valve 1 Feedback - Closed" AND NOT "FPT Tank Vent Valve 1 Feedback - Opened";
END_REGION

REGION Network 5: I0.4 - Tank Vent Valve 2 Feedback Open (CV-441-B)
   // True = OPEN, False = NOT
   RUNG wire#powerrail
      Contact( "FPT Tank Vent Valve 2 Feedback - Opened" )
      I_Contact( "FPT Tank Vent Valve 2 Feedback - Closed" )
      Coil( "20_TANKS_IP_DATA".RIO_01.FIRST_TANK.TANK_VENT_B_OPEN )
   END_RUNG
   // the same network as SCL:
   "20_TANKS_IP_DATA".RIO_01.FIRST_TANK.TANK_VENT_B_OPEN := "FPT Tank Vent Valve 2 Feedback - Opened" AND NOT "FPT Tank Vent Valve 2 Feedback - Closed";
END_REGION

REGION Network 6: I0.5 - Tank Vent Valve 2 Feedback Closed (CV-441-B)
   // True = CLOSED, False = NOT
   RUNG wire#powerrail
      Contact( "FPT Tank Vent Valve 2 Feedback - Closed" )
      I_Contact( "FPT Tank Vent Valve 2 Feedback - Opened" )
      Coil( "20_TANKS_IP_DATA".RIO_01.FIRST_TANK.TANK_VENT_B_CLSD )
   END_RUNG
   // the same network as SCL:
   "20_TANKS_IP_DATA".RIO_01.FIRST_TANK.TANK_VENT_B_CLSD := "FPT Tank Vent Valve 2 Feedback - Closed" AND NOT "FPT Tank Vent Valve 2 Feedback - Opened";
END_REGION

REGION Network 7: I0.6 - Spare Input Accesed from Warning FC
   // True = N/A, False = N/A
END_REGION

REGION Network 8: I0.7 - Spare Input
   // True = N/A, False = N/A
   RUNG wire#powerrail
      Contact( "RIO1_SPR_DI_0_7" )
      Coil( "20_TANKS_IP_DATA".RIO_01.FIRST_TANK.SPARE_DI_7 )
   END_RUNG
   // the same network as SCL:
   "20_TANKS_IP_DATA".RIO_01.FIRST_TANK.SPARE_DI_7 := "RIO1_SPR_DI_0_7";
END_REGION

REGION Network 9: I3.0 - Gas To Tank Valve Feedback Open (CV-422)
   // True = OPEN, False = NOT
   RUNG wire#powerrail
      Contact( "Tank 1P GTT Isolation Valve Feedback - Opened" )
      I_Contact( "Tank 1P GTT Isolation Valve Feedback - Closed" )
      Coil( "20_TANKS_IP_DATA".RIO_01.SECOND_TANK.GTT_ISOL_VALVE_OPEN )
   END_RUNG
   // the same network as SCL:
   "20_TANKS_IP_DATA".RIO_01.SECOND_TANK.GTT_ISOL_VALVE_OPEN := "Tank 1P GTT Isolation Valve Feedback - Opened" AND NOT "Tank 1P GTT Isolation Valve Feedback - Closed";
END_REGION

REGION Network 10: I3.1 - Gas To Tank Valve Feedback Closed (CV-422)
   // True = CLOSED, False = NOT